(* Logix 5000 project; controller _GigaDiscovery vendor 1 type 14 code 244 rev 35.11; software revision 35.03; part 7 of 23 *)
(* tags used below, declared in another part *)
   I_OCC2_Stop_Cycle_PB_memory : BOOL;
   O_Lapbars_Open : ALIAS FOR K300_OCC:5:O.4;
   Output_Scalaggi : Scale_2_P[16];
   SFQ_disable : BOOL;
   SFQ_Mask : DINT;
   SFQ_MASK_OK : DINT;
   Acc_Time : REAL;   // T2 Region 2
   Analog_Output_Pos_5 : REAL[8];
   Angle_at_Full_Load : REAL;
   Angle_at_min_Load : REAL;
   Angle_Controll_S_Curve : S_Curve_Calc;
   auto_manual : TIMER;
   Clock : DINT;   // Base tempi 10 milli sec
   Clock_1_Hz : BOOL;   // SL Clock 1 Hz 0.5 sec OFF 0.5 sec ON
   Clock_4_Hz : BOOL;   // SL Clock 4 Hz 0.125 sec OFF 0.125 sec ON
   Cycle_Time : TIMER;
   First_Push_Set_Torque_to_Zero : BOOL;
   Flyng_Start_Req : BOOL;
   Gate_Entry_Unlock_Selector : BOOL;   // -S30701F
   Gondola_Speed_Reference : DINT;
   Gondola_Torque_Lim : REAL;
   HMI_Horn_Pb : BOOL;   // HMIN Horn Pushbutton
   HMI_Lamp_Test : BOOL;
   HMI_Pylon_Start_Delay : DINT;
   I_EStop_Pb_OCC1 : UDT_DCI_STOP_TEST;   // +OCC E-stop -S30301F
   I_EStop_Pb_OCC2 : UDT_DCI_STOP_TEST;   // +OCC2 E-Stop -S28502F
   I_Fire_Interface : UDT_DCM;   // Page 44
   I_Light_Selector : BOOL;   // Light Selector Switch -S30408F
   I_OCC1_Stop_Cycle_PB : BOOL;   // Stop Cycle -S30308F
   I_OCC2_Disable : UDT_DCM;   // OCC 2 CONTROL DISABLE Page 310
   I_OCC2_Stop_Cycle_PB : BOOL;   // Stop Cycle -S28606F
   I_OCC_Memory_Footpedal : BOOL;
   I_Start_PB : Start_AOI;   // Primary console Strat Push botton Right and Left -S30401F -S30403F
   Jerk_Time : REAL;   // T1 Region 1
   K_Inversion : REAL;   // Fattore di Inversione
   LPF_WLang_Speed_to_Torq : REAL;
   Maintenance_mode : BOOL;   // Ciclo manutenzione per rotazione girella
   Max_Empty_Torque : REAL;   // 75
   Max_Full_Torque : REAL;   // 85
   Mem_RESTRAINTS_closed_Correctly : BOOL;
   Min_Torque_to_Maintain_Height_Full_Load : REAL;
   Min_Torque_to_Maintain_Height_min_Load : REAL;
   MODE : BOOL;   // MODE 0 = AUTO 1 = MANUAL -S30801F
   No_Automatic_E_Stop_Cl_0_Request : BOOL;
   No_Automatic_E_Stop_Cl_1_Request : BOOL;
   No_Emergencies_CL0 : BOOL;
   No_Emergencies_CL1 : BOOL;
   No_Sfty : Std_to_Sfty;
   O_Front_Leg_Light : BOOL;   // Fron leg and front light signal -K3204H
   O_Gondola_Pendolum_Light : BOOL;   // Gondola and pendulum light signal -K3206H
   O_OCC2_Alarms_Lamp : BOOL;
   O_OCC2_Alarms_Noise : BOOL;
   O_Rear_Leg_Light : BOOL;   // Rear leg and rear light signal -K3202H
   O_Sl_RESTRAINTS_Close : ALIAS FOR K300_OCC:5:O.3;
   Os_to_CW_CCW : BOOL;
   Oscillation_Phase : BOOL;
   Platform_Open_Cycle : Sequencer;
   pulse_2_sec : TIMER;
   Pylon_Axe : Axe;
   Pylon_Home_Position : UDT_DCM;   // Home position Pylon -B26002I -B26007I
   Pylon_Seq_Std : Sequencer_AOI_Std;
   Pylon_Speed_Ref : DINT;
   Pylon_Stop_Phase : BOOL;
   Pylon_Stopped_At_Home : BOOL;   // 5s
   Pylon_Torque_Limit : DINT;
   Real : REAL[32];
   RESTRAINTS_Closed : BOOL;   // All RESTRAINTS Closed
   Restraints_Cycle : Sequencer;
   Restraints_Permissive : Permissive;
   RESTRAINTS_Sector : LapBars_Sector[9];
   SCP_K : STD_SCP;
   SCuve_K_Stop : S_Curve_Calc;
   Second_Oscillation_Done : BOOL;   // Second Oscillation End
   Speed_Treshold : REAL;
   Start_Permissive : Permissive;
   Start_Platform_AutoCycle_Pylon : BOOL;
   Start_Stop_Cycle : Sequencer;
   Stop_K_to_Zero : BOOL;
   Stop_Request : BOOL;
   Target_Angle : REAL;
   Timers : TIMER[32];
   To_Sfty : Std_to_Sfty;
   Torque_Filter : REAL;
   Torque_To_Zero_Stewp_04 : BOOL;
   Work_Auto_Cycle_Ptr : DINT;
(* Output, continued *)

ROUTINE _02_Secondary_OCC   (* ladder *)
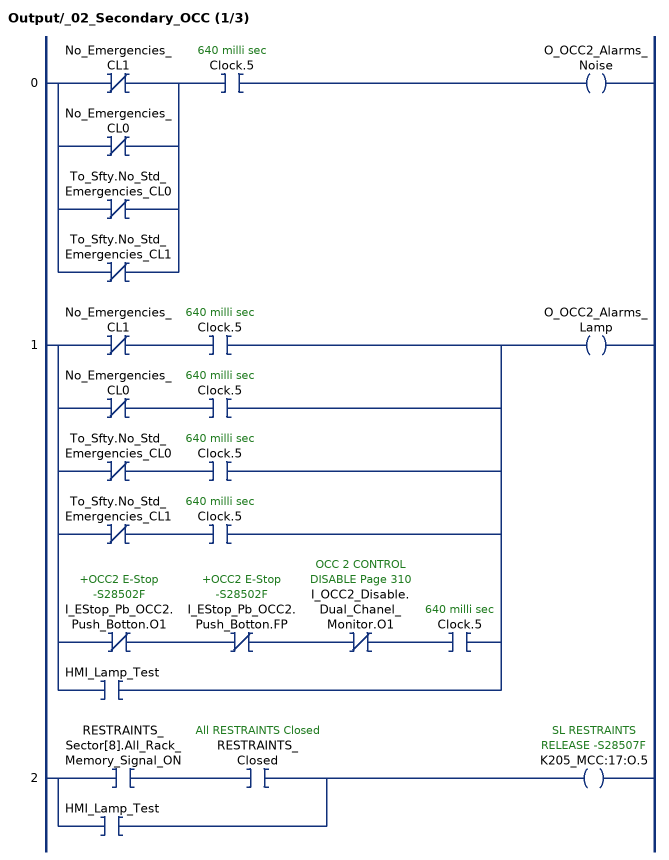
   0: [XIO(No_Emergencies_CL1) ,XIO(No_Emergencies_CL0) ,XIO(To_Sfty.No_Std_Emergencies_CL0) ,XIO(To_Sfty.No_Std_Emergencies_CL1) ]XIC(Clock.5)OTE(O_OCC2_Alarms_Noise);
   1: [XIO(No_Emergencies_CL1) XIC(Clock.5) ,XIO(No_Emergencies_CL0) XIC(Clock.5) ,XIO(To_Sfty.No_Std_Emergencies_CL0) XIC(Clock.5) ,XIO(To_Sfty.No_Std_Emergencies_CL1) XIC(Clock.5) ,XIO(I_EStop_Pb_OCC2.Push_Botton.O1) XIO(I_EStop_Pb_OCC2.Push_Botton.FP) XIO(I_OCC2_Disable.Dual_Chanel_Monitor.O1) XIC(Clock.5) ,XIC(HMI_Lamp_Test) ]OTE(O_OCC2_Alarms_Lamp);
   2: [XIC(RESTRAINTS_Sector[8].All_Rack_Memory_Signal_ON) XIC(RESTRAINTS_Closed) ,XIC(HMI_Lamp_Test) ]OTE(K205_MCC:17:O.5);
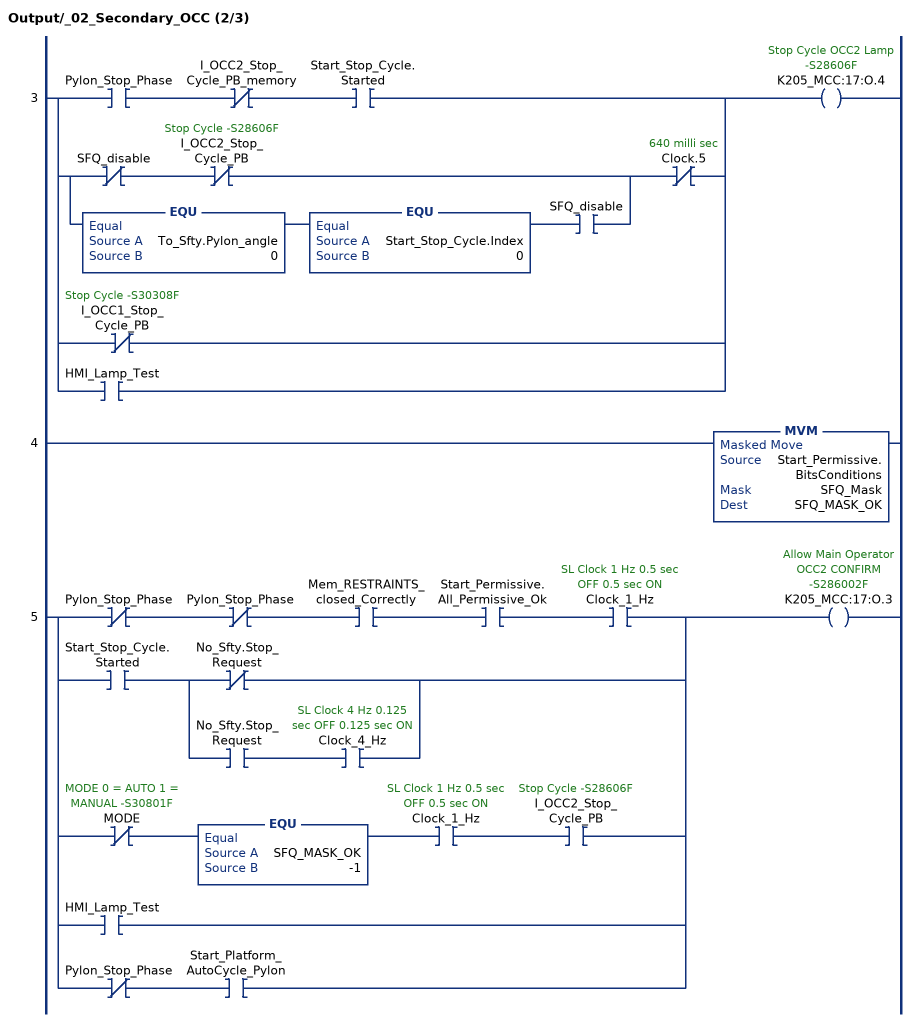
   3: [XIC(Pylon_Stop_Phase) XIO(I_OCC2_Stop_Cycle_PB_memory) XIC(Start_Stop_Cycle.Started) ,[XIO(SFQ_disable) XIO(I_OCC2_Stop_Cycle_PB) ,EQU(To_Sfty.Pylon_angle,0) EQU(Start_Stop_Cycle.Index,0) XIC(SFQ_disable) ] XIO(Clock.5) ,XIO(I_OCC1_Stop_Cycle_PB) ,XIC(HMI_Lamp_Test) ]OTE(K205_MCC:17:O.4);
   4: MVM(Start_Permissive.BitsConditions,SFQ_Mask,SFQ_MASK_OK);
   5: [[XIO(Pylon_Stop_Phase) XIO(Pylon_Stop_Phase) XIC(Mem_RESTRAINTS_closed_Correctly) XIC(Start_Permissive.All_Permissive_Ok) XIC(Clock_1_Hz) ,XIC(Start_Stop_Cycle.Started) [XIO(No_Sfty.Stop_Request) ,XIC(No_Sfty.Stop_Request) XIC(Clock_4_Hz) ] ] ,XIO(MODE) EQU(SFQ_MASK_OK,-1) XIC(Clock_1_Hz) XIC(I_OCC2_Stop_Cycle_PB) ,XIC(HMI_Lamp_Test) ,XIO(Pylon_Stop_Phase) XIC(Start_Platform_AutoCycle_Pylon) ]OTE(K205_MCC:17:O.3);
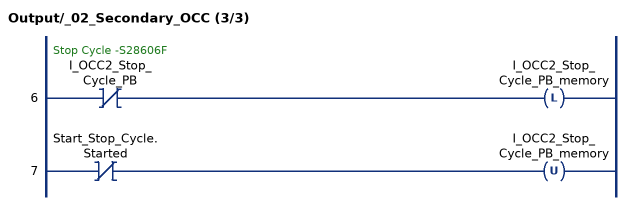
   6: XIO(I_OCC2_Stop_Cycle_PB)OTL(I_OCC2_Stop_Cycle_PB_memory);
   7: XIO(Start_Stop_Cycle.Started)OTU(I_OCC2_Stop_Cycle_PB_memory);
END_ROUTINE

ROUTINE _03_MCC   (* ladder *)
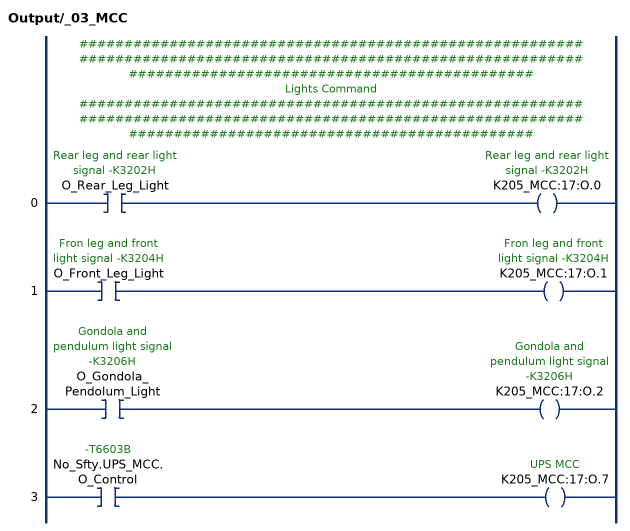
   // #############################################################################################################################################################
   // Lights Command
   // #############################################################################################################################################################
   0: XIC(O_Rear_Leg_Light)OTE(K205_MCC:17:O.0);
   1: XIC(O_Front_Leg_Light)OTE(K205_MCC:17:O.1);
   2: XIC(O_Gondola_Pendolum_Light)OTE(K205_MCC:17:O.2);
   3: XIC(No_Sfty.UPS_MCC.O_Control)OTE(K205_MCC:17:O.7);
END_ROUTINE

ROUTINE _04_RESTRAINTS   (* ladder *)
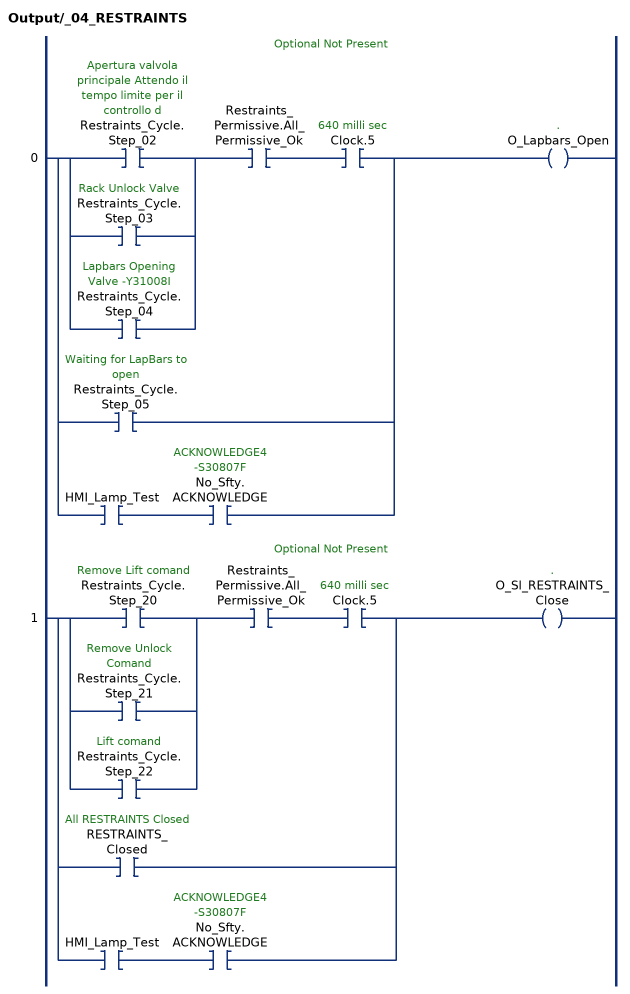
   // Optional Not Present
   0: [[XIC(Restraints_Cycle.Step_02) ,XIC(Restraints_Cycle.Step_03) ,XIC(Restraints_Cycle.Step_04) ] XIC(Restraints_Permissive.All_Permissive_Ok) XIC(Clock.5) ,XIC(Restraints_Cycle.Step_05) ,XIC(HMI_Lamp_Test) XIC(No_Sfty.ACKNOWLEDGE) ]OTE(O_Lapbars_Open);
   // Optional Not Present
   1: [[XIC(Restraints_Cycle.Step_20) ,XIC(Restraints_Cycle.Step_21) ,XIC(Restraints_Cycle.Step_22) ] XIC(Restraints_Permissive.All_Permissive_Ok) XIC(Clock.5) ,XIC(RESTRAINTS_Closed) ,XIC(HMI_Lamp_Test) XIC(No_Sfty.ACKNOWLEDGE) ]OTE(O_Sl_RESTRAINTS_Close);
END_ROUTINE

ROUTINE _06_RCC_02   (* ladder *)
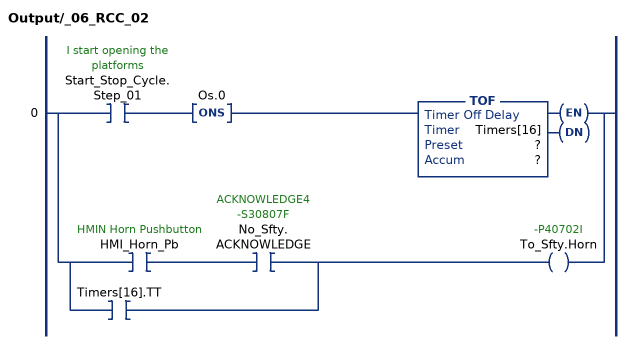
   0: [XIC(Start_Stop_Cycle.Step_01) ONS(Os.0) TOF(Timers[16],?,?) ,[XIC(HMI_Horn_Pb) XIC(No_Sfty.ACKNOWLEDGE) ,XIC(Timers[16].TT) ] OTE(To_Sfty.Horn) ];
END_ROUTINE

ROUTINE _07_External_Interface   (* ladder *)
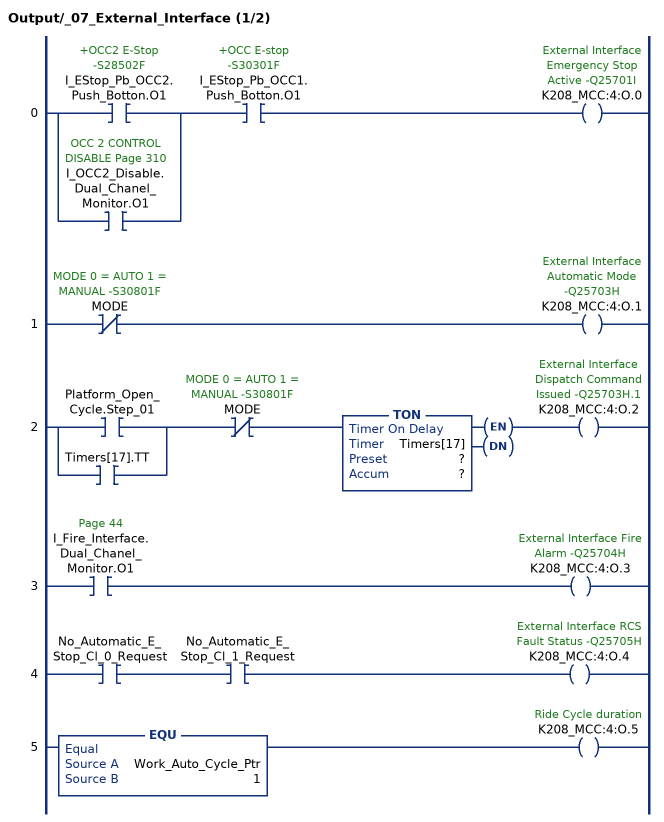
   0: [XIC(I_EStop_Pb_OCC2.Push_Botton.O1) ,XIC(I_OCC2_Disable.Dual_Chanel_Monitor.O1) ]XIC(I_EStop_Pb_OCC1.Push_Botton.O1)OTE(K208_MCC:4:O.0);
   1: XIO(MODE)OTE(K208_MCC:4:O.1);
   2: [XIC(Platform_Open_Cycle.Step_01) ,XIC(Timers[17].TT) ]XIO(MODE)TON(Timers[17],?,?)OTE(K208_MCC:4:O.2);
   3: XIC(I_Fire_Interface.Dual_Chanel_Monitor.O1)OTE(K208_MCC:4:O.3);
   4: XIC(No_Automatic_E_Stop_Cl_0_Request)XIC(No_Automatic_E_Stop_Cl_1_Request)OTE(K208_MCC:4:O.4);
   5: EQU(Work_Auto_Cycle_Ptr,1)OTE(K208_MCC:4:O.5);
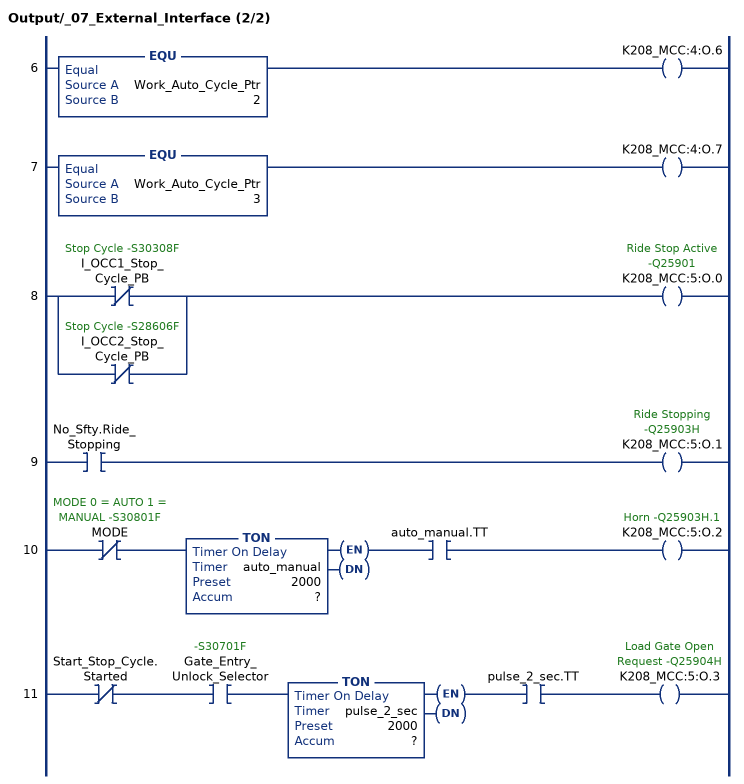
   6: EQU(Work_Auto_Cycle_Ptr,2)OTE(K208_MCC:4:O.6);
   7: EQU(Work_Auto_Cycle_Ptr,3)OTE(K208_MCC:4:O.7);
   8: [XIO(I_OCC1_Stop_Cycle_PB) ,XIO(I_OCC2_Stop_Cycle_PB) ]OTE(K208_MCC:5:O.0);
   9: XIC(No_Sfty.Ride_Stopping)OTE(K208_MCC:5:O.1);
   10: XIO(MODE)TON(auto_manual,?,?)XIC(auto_manual.TT)OTE(K208_MCC:5:O.2);
   11: XIO(Start_Stop_Cycle.Started)XIC(Gate_Entry_Unlock_Selector)TON(pulse_2_sec,?,?)XIC(pulse_2_sec.TT)OTE(K208_MCC:5:O.3);
END_ROUTINE

ROUTINE Main   (* ladder *)
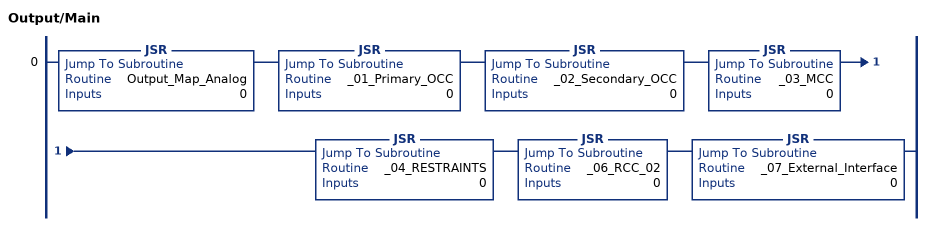
   0: JSR(Output_Map_Analog,0)JSR(_01_Primary_OCC,0)JSR(_02_Secondary_OCC,0)JSR(_03_MCC,0)JSR(_04_RESTRAINTS,0)JSR(_06_RCC_02,0)JSR(_07_External_Interface,0);
END_ROUTINE

ROUTINE Output_Map_Analog   (* function block diagram *)
   SHEET 1   // Pilon
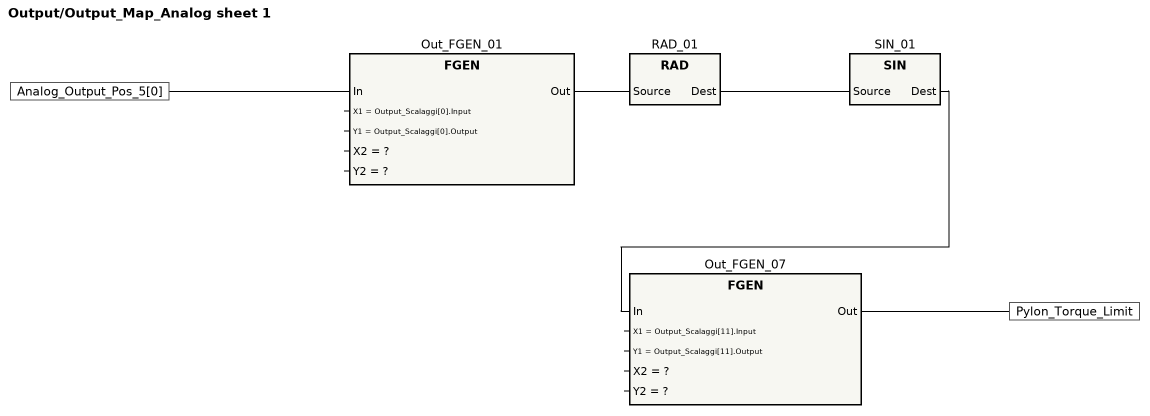
   Out_FGEN_01 : FGEN(In := Analog_Output_Pos_5[0], X1 := Output_Scalaggi[0].Input, Y1 := Output_Scalaggi[0].Output, X2 := ?, Y2 := ?);
   RAD_01 : RAD(Source := Out_FGEN_01.Out);
   SIN_01 : SIN(Source := RAD_01.Dest);
   Out_FGEN_07 : FGEN(In := SIN_01.Dest, X1 := Output_Scalaggi[11].Input, Y1 := Output_Scalaggi[11].Output, X2 := ?, Y2 := ?);
   Pylon_Torque_Limit := Out_FGEN_07.Out;
   SHEET 2   // Gondola
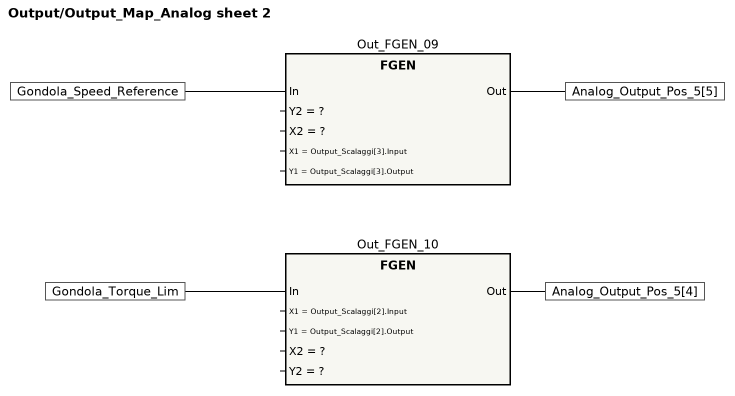
   Out_FGEN_09 : FGEN(In := Gondola_Speed_Reference, Y2 := ?, X2 := ?, X1 := Output_Scalaggi[3].Input, Y1 := Output_Scalaggi[3].Output);
   Out_FGEN_10 : FGEN(In := Gondola_Torque_Lim, X1 := Output_Scalaggi[2].Input, Y1 := Output_Scalaggi[2].Output, X2 := ?, Y2 := ?);
   Analog_Output_Pos_5[4] := Out_FGEN_10.Out;
   Analog_Output_Pos_5[5] := Out_FGEN_09.Out;
   SHEET 3   // Gondola V and I
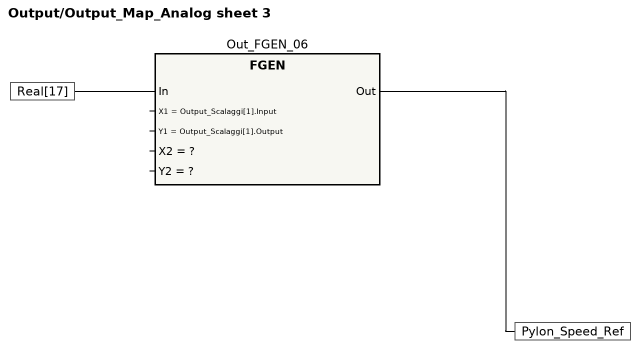
   Out_FGEN_06 : FGEN(In := Real[17], X1 := Output_Scalaggi[1].Input, Y1 := Output_Scalaggi[1].Output, X2 := ?, Y2 := ?);
   Pylon_Speed_Ref := Out_FGEN_06.Out;
END_ROUTINE
END_PROGRAM

PROGRAM Pylon   (* main routine Main *)
VAR
   ArmInductanceGondola : REAL := 5.494;
   ArmResistanceGondola : REAL := 0.49;
   First_Push_Angle : REAL := 13.991667;   // WEIGHT
   Gondola_Start_Delay : TIMER := (PRE := 5000);
   Gondola_Stop : BOOL;
   JM_ons : DINT;
   JM_RunEnd : TIMER := (PRE := 240000);
   K_Edge_Push_Up : DINT[10] := ([0] := 30, [1] := 50, [2] := 80);
   Max_Torque_for_Angle_Correction : REAL := 84.066666;
   Min_error_to_Start_Decreasing_Torque : REAL := 10.0;
   Os : DINT := 384;
   Os_to_CCW : BOOL;
   Os_to_CW : BOOL;
   Pylon_Real : REAL[10] := ([0] := 1.0, [1] := 5.0, [2] := 18.0, [3] := 0.1, [4] := 5.0);
   Pylon_Sequencer : Sequencer := (Step_Timer[0].PRE := 100, Step_Timer[1].PRE := 4000, Step_Timer[2].PRE := 250, Step_Timer[3].PRE := 4000, Step_Timer[4].PRE := 1250, Step_Timer[5].PRE := 2000, Step_Timer[31].PRE := 7500, Step_Timer[31].ACC := 7500, Step_Timer[31].EN := 1, Step_Timer[31].DN := 1, Step_00 := 1);
        .Step_Timer[1]   // Dopo un temp t tolgo coppia per far scendere il pendolo
        .Step_02   // Prima Spinta CCW Calcolo Peso
        .Step_04   // Stop Request
        .Step_03   // Oscillazioni
        .Step_01   // Prima Spinta CW
        .Step_06   // Stop Pilone
        .Step_05   // Quando sono a velocità Bassa Resetto la Posizione
   Pylon_Start_Delay : TIMER;
   RunEndDetails : DINT[10] := ([1] := 107, [2] := 3217, [3] := 71013, [4] := 85950);
        [2]   // time at step 5
        [1]   // last angle
        [4]   // time at step 6 end
        [3]   // time at step 6
   SCL_01_Loc1 : SCALE := (In := 13.991667, InRawMax := 14.0, InRawMin := 12.0, InEUMax := 84.0, InEUMin := 100.0, Limiting := 1, Out := 84.066666);
   SCL_01_Loc1_01 : SCALE := (In := 8.841667, InRawMax := 10.0, InRawMin := -2.0, InEUMax := 84.066666, InEUMin := 15.0, Limiting := 1, Out := 77.39982);
   SCL_01_Loc1_02 : SCALE := (In := 13.991667, InRawMax := 14.0, InRawMin := 12.0, InEUMax := 15.0, InEUMin := 15.0, Limiting := 1, Out := 15.0);
   SpeedRegKi : REAL := 20.0;
   SpeedRegKp : REAL := 10.0;
   Timer : TIMER[10] := ([0].PRE := 9500, [1].PRE := 1000, [2].PRE := 100, [3].PRE := 5500, [4].PRE := 6500, [5].PRE := 7000);
END_VAR

ROUTINE _00_Settings   (* ladder *)
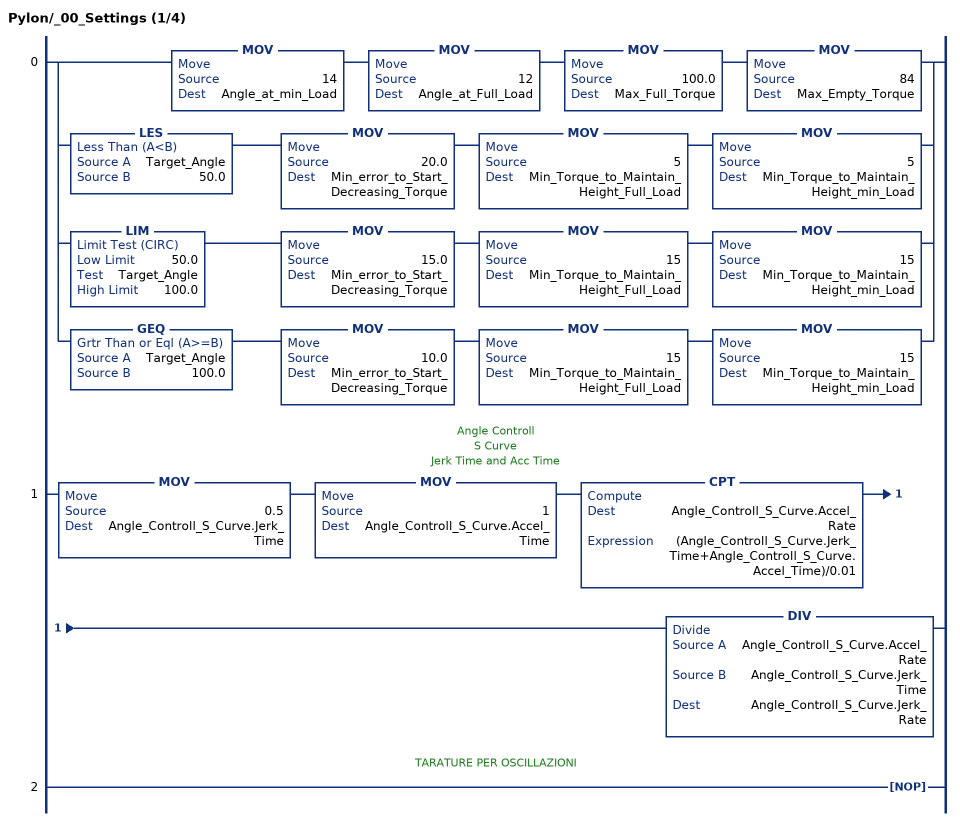
   0: [MOV(14,Angle_at_min_Load) MOV(12,Angle_at_Full_Load) MOV(100.0,Max_Full_Torque) MOV(84,Max_Empty_Torque) ,LES(Target_Angle,50.0) MOV(20.0,Min_error_to_Start_Decreasing_Torque) MOV(5,Min_Torque_to_Maintain_Height_Full_Load) MOV(5,Min_Torque_to_Maintain_Height_min_Load) ,LIM(50.0,Target_Angle,100.0) MOV(15.0,Min_error_to_Start_Decreasing_Torque) MOV(15,Min_Torque_to_Maintain_Height_Full_Load) MOV(15,Min_Torque_to_Maintain_Height_min_Load) ,GEQ(Target_Angle,100.0) MOV(10.0,Min_error_to_Start_Decreasing_Torque) MOV(15,Min_Torque_to_Maintain_Height_Full_Load) MOV(15,Min_Torque_to_Maintain_Height_min_Load) ];
   // Angle Controll
   // S Curve
   // Jerk Time and Acc Time
   1: MOV(0.5,Angle_Controll_S_Curve.Jerk_Time)MOV(1,Angle_Controll_S_Curve.Accel_Time)CPT(Angle_Controll_S_Curve.Accel_Rate,(Angle_Controll_S_Curve.Jerk_Time+Angle_Controll_S_Curve.Accel_Time)/0.01)DIV(Angle_Controll_S_Curve.Accel_Rate,Angle_Controll_S_Curve.Jerk_Time,Angle_Controll_S_Curve.Jerk_Rate);
   // TARATURE PER OSCILLAZIONI
   2: NOP();
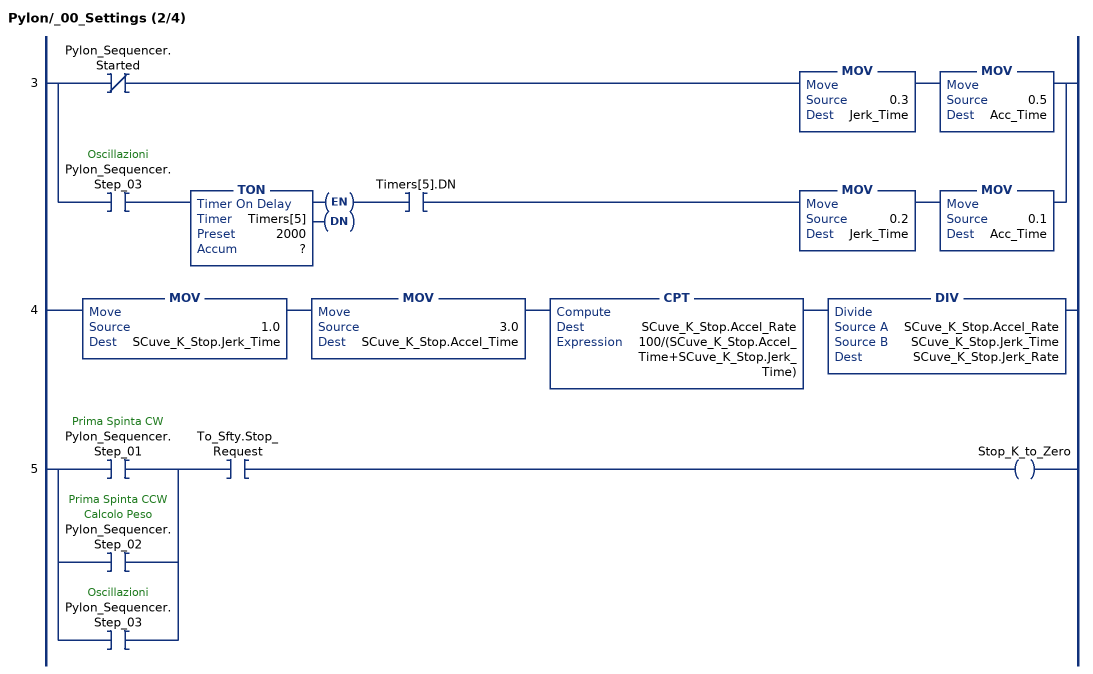
   3: [XIO(Pylon_Sequencer.Started) MOV(0.3,Jerk_Time) MOV(0.5,Acc_Time) ,XIC(Pylon_Sequencer.Step_03) TON(Timers[5],?,?) XIC(Timers[5].DN) MOV(0.2,Jerk_Time) MOV(0.1,Acc_Time) ];
   4: MOV(1.0,SCuve_K_Stop.Jerk_Time)MOV(3.0,SCuve_K_Stop.Accel_Time)CPT(SCuve_K_Stop.Accel_Rate,100/(SCuve_K_Stop.Accel_Time+SCuve_K_Stop.Jerk_Time))DIV(SCuve_K_Stop.Accel_Rate,SCuve_K_Stop.Jerk_Time,SCuve_K_Stop.Jerk_Rate);
   5: [XIC(Pylon_Sequencer.Step_01) ,XIC(Pylon_Sequencer.Step_02) ,XIC(Pylon_Sequencer.Step_03) ]XIC(To_Sfty.Stop_Request)OTE(Stop_K_to_Zero);
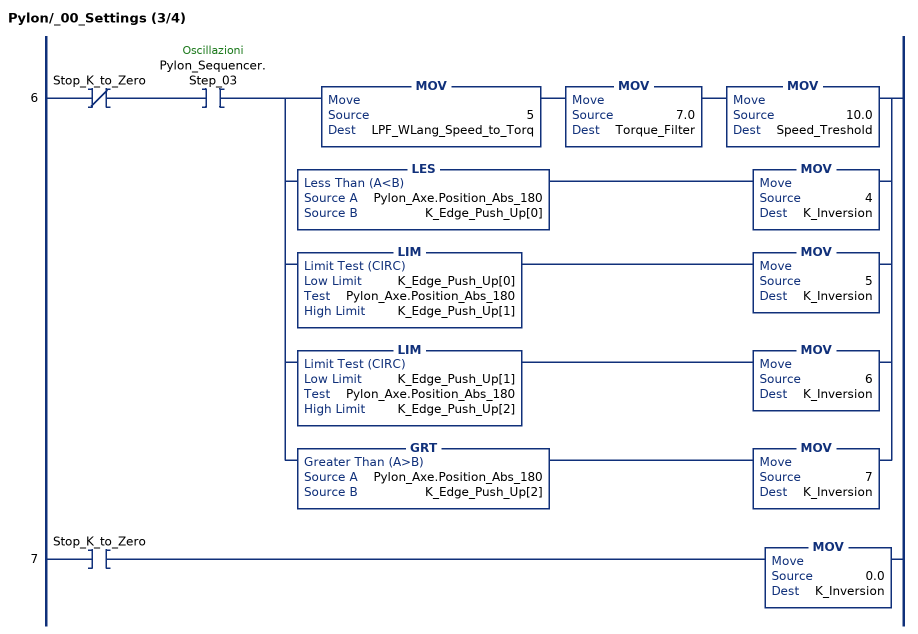
   6: XIO(Stop_K_to_Zero)XIC(Pylon_Sequencer.Step_03)[MOV(5,LPF_WLang_Speed_to_Torq) MOV(7.0,Torque_Filter) MOV(10.0,Speed_Treshold) ,LES(Pylon_Axe.Position_Abs_180,K_Edge_Push_Up[0]) MOV(4,K_Inversion) ,LIM(K_Edge_Push_Up[0],Pylon_Axe.Position_Abs_180,K_Edge_Push_Up[1]) MOV(5,K_Inversion) ,LIM(K_Edge_Push_Up[1],Pylon_Axe.Position_Abs_180,K_Edge_Push_Up[2]) MOV(6,K_Inversion) ,GRT(Pylon_Axe.Position_Abs_180,K_Edge_Push_Up[2]) MOV(7,K_Inversion) ];
   7: XIC(Stop_K_to_Zero)MOV(0.0,K_Inversion);
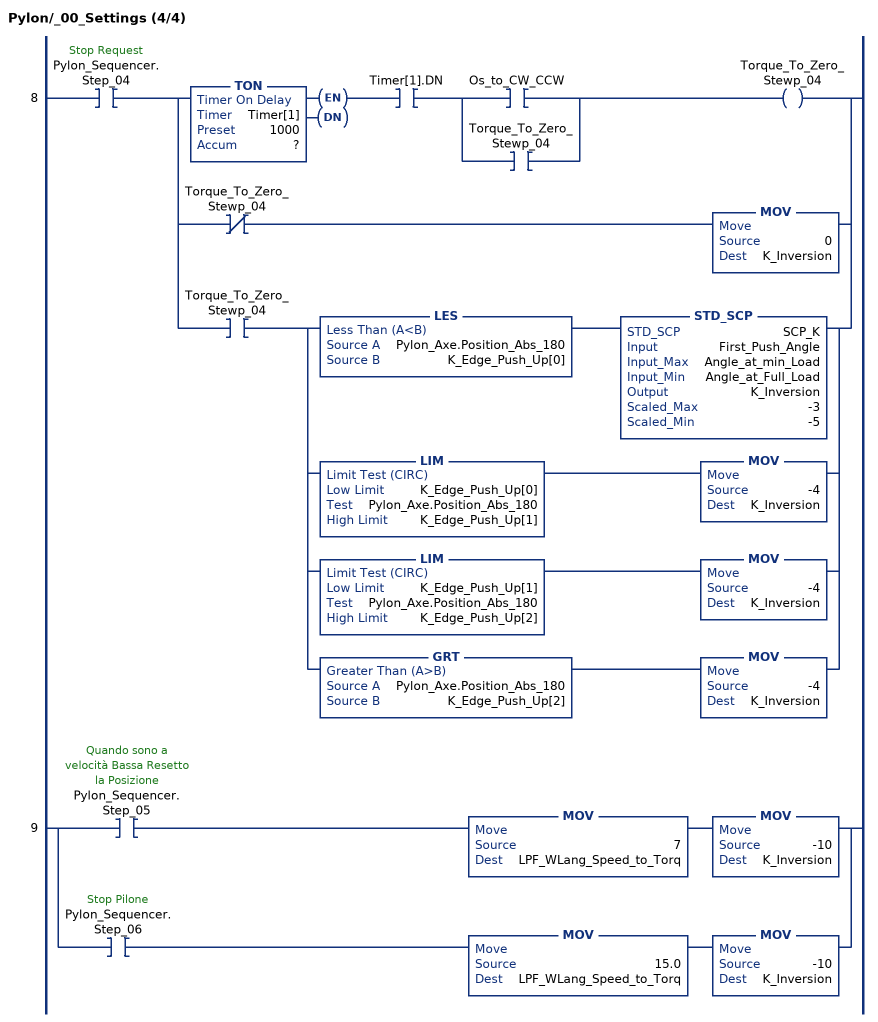
   8: XIC(Pylon_Sequencer.Step_04)[TON(Timer[1],?,?) XIC(Timer[1].DN) [XIC(Os_to_CW_CCW) ,XIC(Torque_To_Zero_Stewp_04) ] OTE(Torque_To_Zero_Stewp_04) ,XIO(Torque_To_Zero_Stewp_04) MOV(0,K_Inversion) ,XIC(Torque_To_Zero_Stewp_04) [LES(Pylon_Axe.Position_Abs_180,K_Edge_Push_Up[0]) STD_SCP(SCP_K,First_Push_Angle,Angle_at_min_Load,Angle_at_Full_Load,K_Inversion,-3,-5) ,LIM(K_Edge_Push_Up[0],Pylon_Axe.Position_Abs_180,K_Edge_Push_Up[1]) MOV(-4,K_Inversion) ,LIM(K_Edge_Push_Up[1],Pylon_Axe.Position_Abs_180,K_Edge_Push_Up[2]) MOV(-4,K_Inversion) ,GRT(Pylon_Axe.Position_Abs_180,K_Edge_Push_Up[2]) MOV(-4,K_Inversion) ] ];
   9: [XIC(Pylon_Sequencer.Step_05) MOV(7,LPF_WLang_Speed_to_Torq) MOV(-10,K_Inversion) ,XIC(Pylon_Sequencer.Step_06) MOV(15.0,LPF_WLang_Speed_to_Torq) MOV(-10,K_Inversion) ];
END_ROUTINE

ROUTINE _01_Auto_Cycle   (* ladder *)
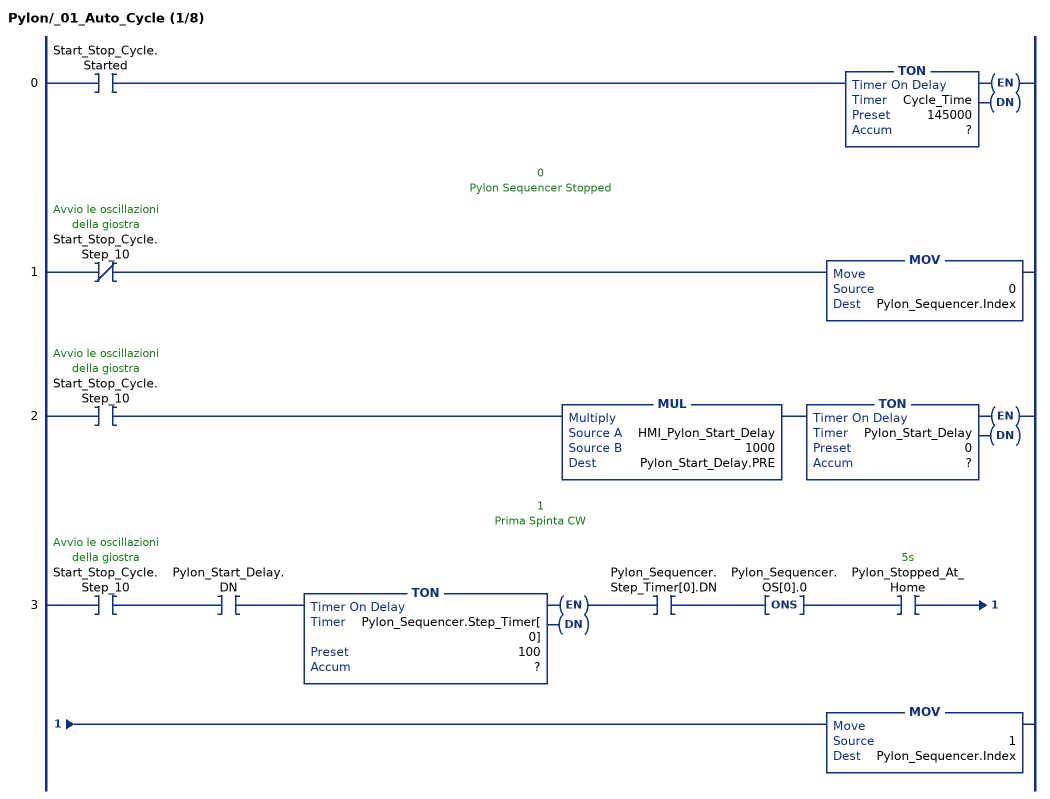
   0: XIC(Start_Stop_Cycle.Started)TON(Cycle_Time,?,?);
   // 0
   // Pylon Sequencer Stopped
   1: XIO(Start_Stop_Cycle.Step_10)MOV(0,Pylon_Sequencer.Index);
   2: XIC(Start_Stop_Cycle.Step_10)MUL(HMI_Pylon_Start_Delay,1000,Pylon_Start_Delay.PRE)TON(Pylon_Start_Delay,?,?);
   // 1
   // Prima Spinta CW
   3: XIC(Start_Stop_Cycle.Step_10)XIC(Pylon_Start_Delay.DN)TON(Pylon_Sequencer.Step_Timer[0],?,?)XIC(Pylon_Sequencer.Step_Timer[0].DN)ONS(Pylon_Sequencer.OS[0].0)XIC(Pylon_Stopped_At_Home)MOV(1,Pylon_Sequencer.Index);
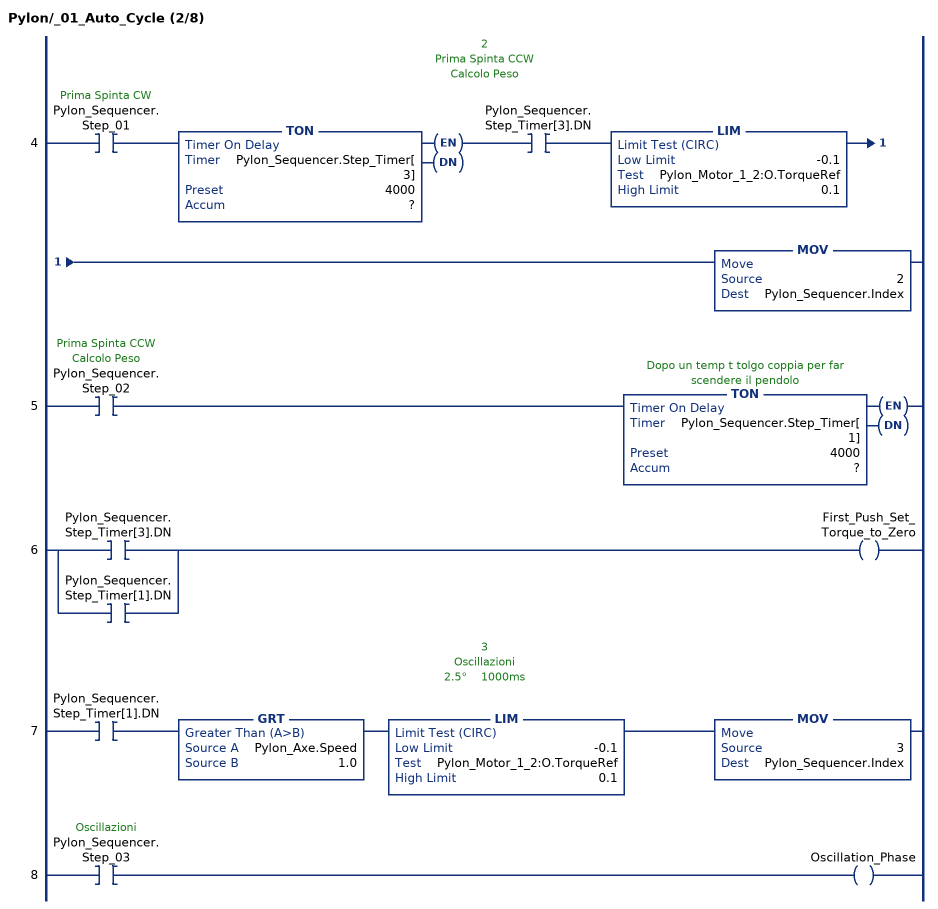
   // 2
   // Prima Spinta CCW
   // Calcolo Peso
   4: XIC(Pylon_Sequencer.Step_01)TON(Pylon_Sequencer.Step_Timer[3],?,?)XIC(Pylon_Sequencer.Step_Timer[3].DN)LIM(-0.1,Pylon_Motor_1_2:O.TorqueRef,0.1)MOV(2,Pylon_Sequencer.Index);
   5: XIC(Pylon_Sequencer.Step_02)TON(Pylon_Sequencer.Step_Timer[1],?,?);
   6: [XIC(Pylon_Sequencer.Step_Timer[3].DN) ,XIC(Pylon_Sequencer.Step_Timer[1].DN) ]OTE(First_Push_Set_Torque_to_Zero);
   // 3
   // Oscillazioni
   // 2.5°    1000ms
   7: XIC(Pylon_Sequencer.Step_Timer[1].DN)GRT(Pylon_Axe.Speed,1.0)LIM(-0.1,Pylon_Motor_1_2:O.TorqueRef,0.1)MOV(3,Pylon_Sequencer.Index);
   8: XIC(Pylon_Sequencer.Step_03)OTE(Oscillation_Phase);
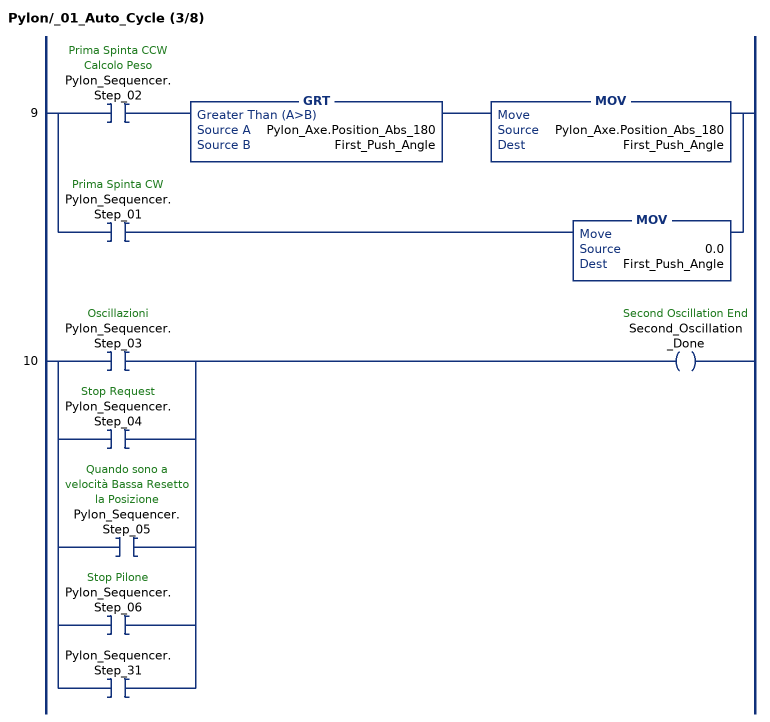
   9: [XIC(Pylon_Sequencer.Step_02) GRT(Pylon_Axe.Position_Abs_180,First_Push_Angle) MOV(Pylon_Axe.Position_Abs_180,First_Push_Angle) ,XIC(Pylon_Sequencer.Step_01) MOV(0.0,First_Push_Angle) ];
   10: [XIC(Pylon_Sequencer.Step_03) ,XIC(Pylon_Sequencer.Step_04) ,XIC(Pylon_Sequencer.Step_05) ,XIC(Pylon_Sequencer.Step_06) ,XIC(Pylon_Sequencer.Step_31) ]OTE(Second_Oscillation_Done);
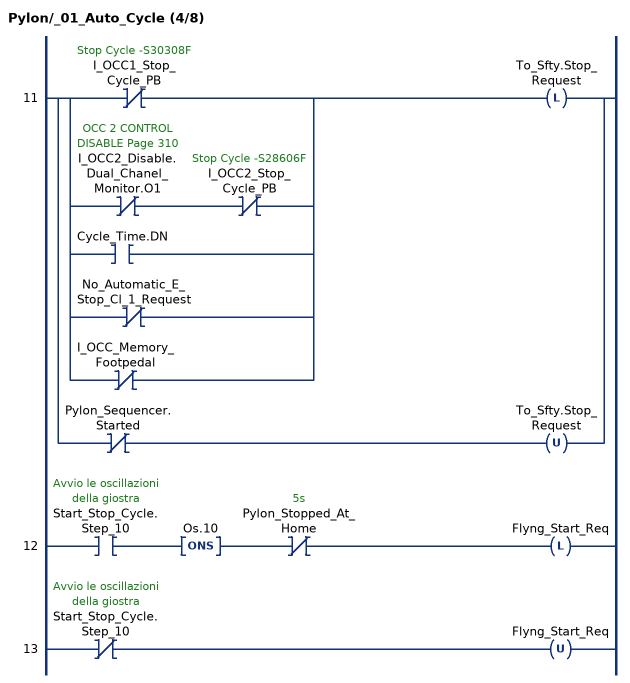
   11: [[XIO(I_OCC1_Stop_Cycle_PB) ,XIO(I_OCC2_Disable.Dual_Chanel_Monitor.O1) XIO(I_OCC2_Stop_Cycle_PB) ,XIC(Cycle_Time.DN) ,XIO(No_Automatic_E_Stop_Cl_1_Request) ,XIO(I_OCC_Memory_Footpedal) ] OTL(To_Sfty.Stop_Request) ,XIO(Pylon_Sequencer.Started) OTU(To_Sfty.Stop_Request) ];
   12: XIC(Start_Stop_Cycle.Step_10)ONS(Os.10)XIO(Pylon_Stopped_At_Home)OTL(Flyng_Start_Req);
   13: XIO(Start_Stop_Cycle.Step_10)OTU(Flyng_Start_Req);
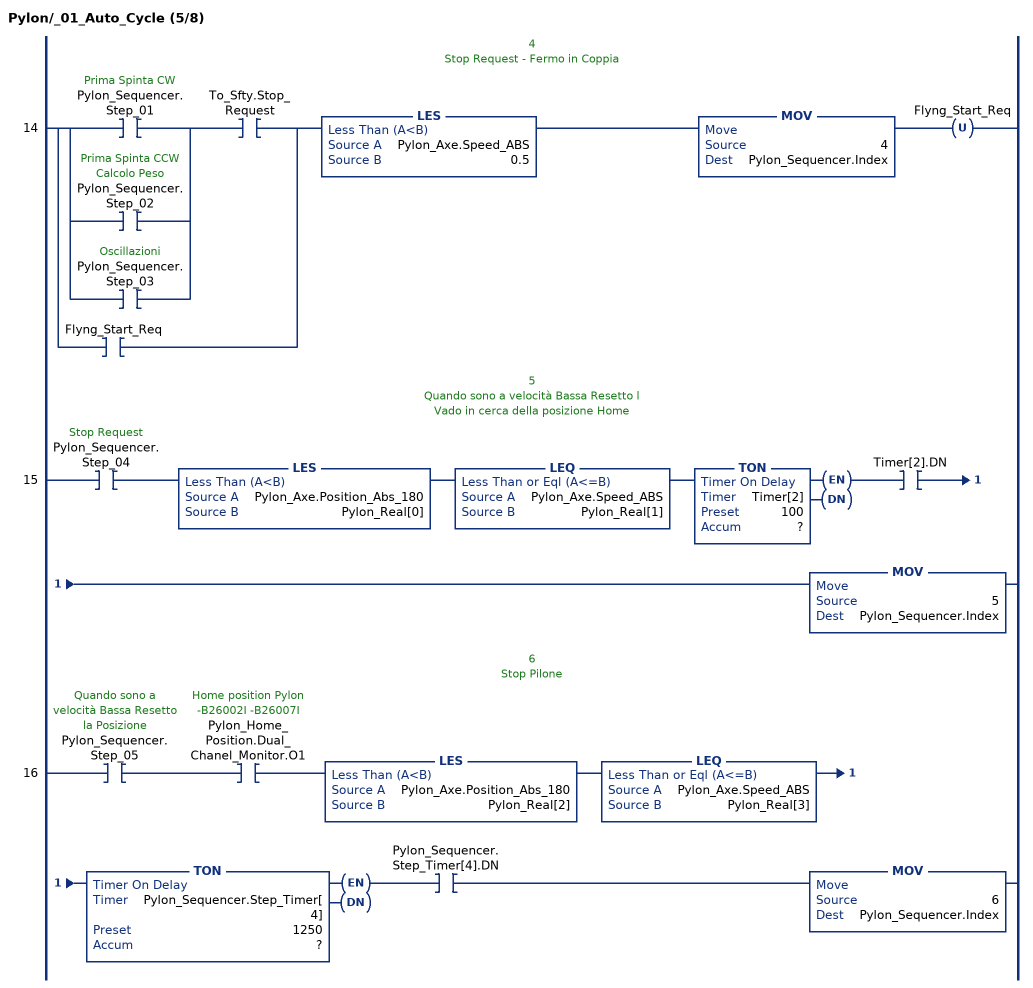
   // 4
   // Stop Request - Fermo in Coppia
   14: [[XIC(Pylon_Sequencer.Step_01) ,XIC(Pylon_Sequencer.Step_02) ,XIC(Pylon_Sequencer.Step_03) ] XIC(To_Sfty.Stop_Request) ,XIC(Flyng_Start_Req) ]LES(Pylon_Axe.Speed_ABS,0.5)MOV(4,Pylon_Sequencer.Index)OTU(Flyng_Start_Req);
   // 5
   // Quando sono a velocità Bassa Resetto l
   // Vado in cerca della posizione Home
   15: XIC(Pylon_Sequencer.Step_04)LES(Pylon_Axe.Position_Abs_180,Pylon_Real[0])LEQ(Pylon_Axe.Speed_ABS,Pylon_Real[1])TON(Timer[2],?,?)XIC(Timer[2].DN)MOV(5,Pylon_Sequencer.Index);
   // 6
   // Stop Pilone
   16: XIC(Pylon_Sequencer.Step_05)XIC(Pylon_Home_Position.Dual_Chanel_Monitor.O1)LES(Pylon_Axe.Position_Abs_180,Pylon_Real[2])LEQ(Pylon_Axe.Speed_ABS,Pylon_Real[3])TON(Pylon_Sequencer.Step_Timer[4],?,?)XIC(Pylon_Sequencer.Step_Timer[4].DN)MOV(6,Pylon_Sequencer.Index);
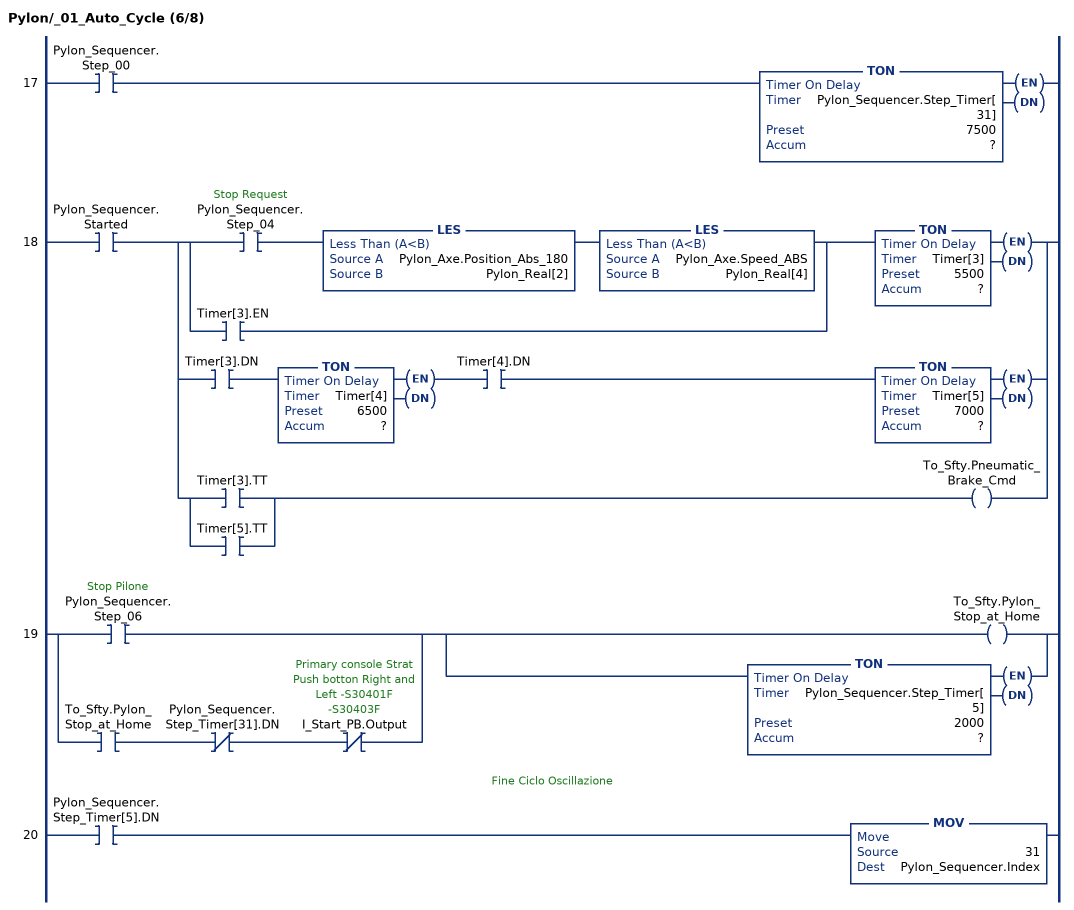
   17: XIC(Pylon_Sequencer.Step_00)TON(Pylon_Sequencer.Step_Timer[31],?,?);
   18: XIC(Pylon_Sequencer.Started)[[XIC(Pylon_Sequencer.Step_04) LES(Pylon_Axe.Position_Abs_180,Pylon_Real[2]) LES(Pylon_Axe.Speed_ABS,Pylon_Real[4]) ,XIC(Timer[3].EN) ] TON(Timer[3],?,?) ,XIC(Timer[3].DN) TON(Timer[4],?,?) XIC(Timer[4].DN) TON(Timer[5],?,?) ,[XIC(Timer[3].TT) ,XIC(Timer[5].TT) ] OTE(To_Sfty.Pneumatic_Brake_Cmd) ];
   19: [XIC(Pylon_Sequencer.Step_06) ,XIC(To_Sfty.Pylon_Stop_at_Home) XIO(Pylon_Sequencer.Step_Timer[31].DN) XIO(I_Start_PB.Output) ][OTE(To_Sfty.Pylon_Stop_at_Home) ,TON(Pylon_Sequencer.Step_Timer[5],?,?) ];
   // Fine Ciclo Oscillazione
   20: XIC(Pylon_Sequencer.Step_Timer[5].DN)MOV(31,Pylon_Sequencer.Index);
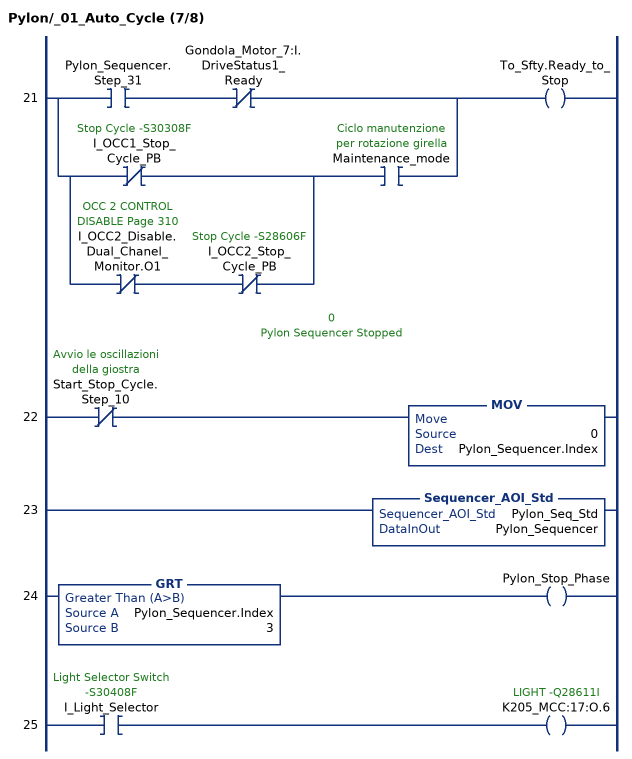
   21: [XIC(Pylon_Sequencer.Step_31) XIO(Gondola_Motor_7:I.DriveStatus1_Ready) ,[XIO(I_OCC1_Stop_Cycle_PB) ,XIO(I_OCC2_Disable.Dual_Chanel_Monitor.O1) XIO(I_OCC2_Stop_Cycle_PB) ] XIC(Maintenance_mode) ]OTE(To_Sfty.Ready_to_Stop);
   // 0
   // Pylon Sequencer Stopped
   22: XIO(Start_Stop_Cycle.Step_10)MOV(0,Pylon_Sequencer.Index);
   23: Sequencer_AOI_Std(Pylon_Seq_Std,Pylon_Sequencer);
   24: GRT(Pylon_Sequencer.Index,3)OTE(Pylon_Stop_Phase);
   25: XIC(I_Light_Selector)OTE(K205_MCC:17:O.6);
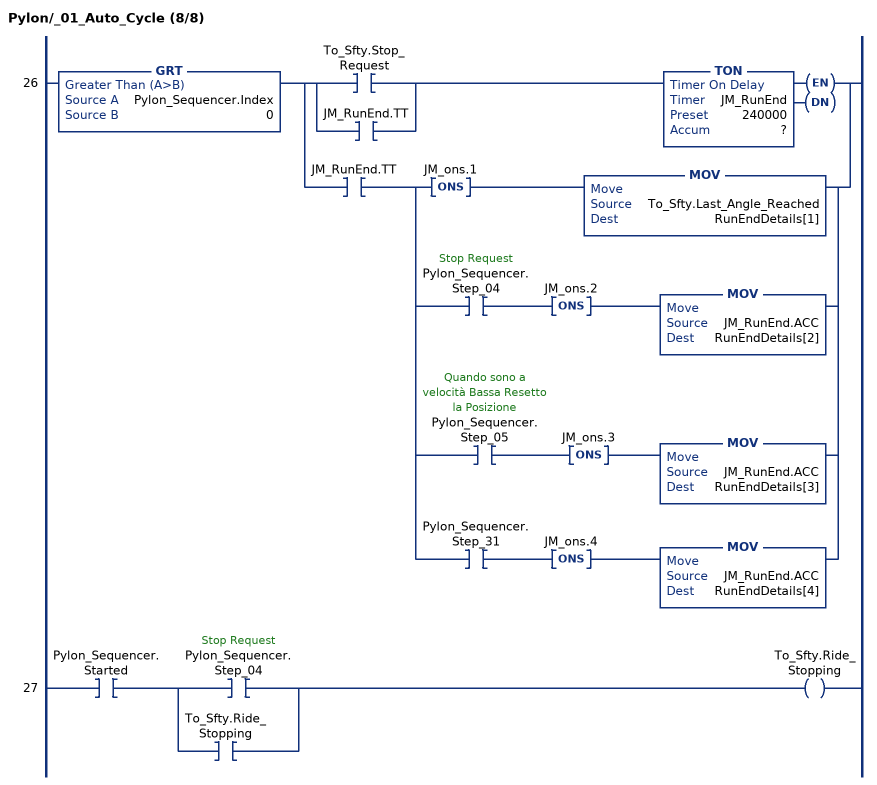
   26: GRT(Pylon_Sequencer.Index,0)[[XIC(To_Sfty.Stop_Request) ,XIC(JM_RunEnd.TT) ] TON(JM_RunEnd,?,?) ,XIC(JM_RunEnd.TT) [ONS(JM_ons.1) MOV(To_Sfty.Last_Angle_Reached,RunEndDetails[1]) ,XIC(Pylon_Sequencer.Step_04) ONS(JM_ons.2) MOV(JM_RunEnd.ACC,RunEndDetails[2]) ,XIC(Pylon_Sequencer.Step_05) ONS(JM_ons.3) MOV(JM_RunEnd.ACC,RunEndDetails[3]) ,XIC(Pylon_Sequencer.Step_31) ONS(JM_ons.4) MOV(JM_RunEnd.ACC,RunEndDetails[4]) ] ];
   27: XIC(Pylon_Sequencer.Started)[XIC(Pylon_Sequencer.Step_04) ,XIC(To_Sfty.Ride_Stopping) ]OTE(To_Sfty.Ride_Stopping);
END_ROUTINE
